(* Logix 5000 project; controller FV vendor 1 type 14 code 217 rev 31.11; software revision 31.00; part 16 of 63 *)
(* tags used below, declared in another part *)
   Dummy : BOOL;
   FR_B230 : INT[255];   // FLOW_BITS Flow Meter Bits
   FR_B240 : INT[255];   // DEBOUNCE Debounce Flags
   FR_B246 : INT[255];   // V_REVERSE Flags for reversing contol action
   FR_B247 : INT[255];   // CHECKWORD Simulation Flags for Checkwords
   FR_B248 : INT[255];   // FORCE ON Force On Flags
   FR_B249 : INT[255];   // FORCE_OFF NOT Force Off Flags
   FR_B3 : INT[255];   // BINARY
   FR_bit_data_file_address : DINT;
   FR_bit_file_bit_offset : DINT;
   FR_bit_file_word_offset : DINT;
   FR_bit_offset : DINT;
   FR_bit_returned : BOOL;
   FR_data_file_value_to_move : DINT;
   FR_from_data_file : DINT;
   FR_from_data_offset : DINT;
   FR_N10 : INT[265];   // FV_AGING Comms to FV Aging PL C
   FR_N100 : INT[265];   // FV FILLING
   FR_N110 : INT[265];   // GREEN BEER Green Beer Main
   FR_N120 : INT[265];   // YEAST CROP Yeast Cropping Main
   FR_N13 : INT[265];   // MV_ROUTE Comms to MV Routing PLC
   FR_N130 : INT[265];   // FILTRATE Filtrate Return
   FR_N14 : INT[265];   // MVFV CIP Comms to MVFV CIP Un it PLC
   FR_N140 : INT[265];   // CIP
   FR_N142 : INT[265];   // CIP
   FR_N143 : INT[265];   // CIP
   FR_N150 : INT[265];   // Original N File From SLC, No Description Available
   FR_N160 : INT[265];   // VESSEL Vessel Working Direc tory
   FR_N170 : INT[265];   // Original N File From SLC, No Description Available
   FR_N180 : INT[265];   // Original N File From SLC, No Description Available
   FR_N198 : INT[265];   // Original N File From SLC, No Description Available
   FR_N20 : INT[265];   // GENERAL General Purpose Setp oints
   FR_N200 : INT[265];   // ANALOG_IN Analog Inputs
   FR_N201 : INT[265];   // Original N File From SLC, No Description Available
   FR_N207 : INT[265];   // Original N File From SLC, No Description Available
   FR_N21 : INT[265];   // CHASE_V FV Filling Beer Chas e Volumes
   FR_N210 : INT[265];   // ANALOG_OUT Analog Outputs
   FR_N220 : INT[265];   // CHECKLIST Checklist Loop Contr ollers
   FR_N225 : INT[265];   // Original N File From SLC, No Description Available
   FR_N226 : INT[265];   // Original N File From SLC, No Description Available
   FR_N245 : INT[265];   // CHECKWORD Checkword Loop Contr ol
   FR_N252 : INT[265];   // OUTPUT_PTR Checkword Pointers t o output flags in B2 50
   FR_N253 : INT[265];   // EN_POINT Pointers to energise d input flags in B25 1
   FR_N254 : INT[265];   // DEN_POINT Pointers to deenergi sed input flags in B 251
   FR_N255 : INT[265];   // CHECKWORDS
   FR_N26 : INT[265];   // FV26
   FR_N27 : INT[265];   // FV27
   FR_N28 : INT[265];   // FV28
   FR_N29 : INT[265];   // FV29
   FR_N30 : INT[265];   // FV30
   FR_N31 : INT[265];   // FV31
   FR_N36 : INT[265];   // Original N File From SLC, No Description Available
   FR_N37 : INT[265];   // Original N File From SLC, No Description Available
   FR_N46 : INT[265];   // Original N File From SLC, No Description Available
   FR_N47 : INT[265];   // Original N File From SLC, No Description Available
   FR_N7 : INT[265];   // INTEGER
   FR_N99 : INT[265];   // COMMENT Comment Lines
   FR_T111 : TIMER[255];   // GREEN BEER
(* FR_Common, continued *)

ROUTINE FR_Get_NFile_Value   (* ladder *)
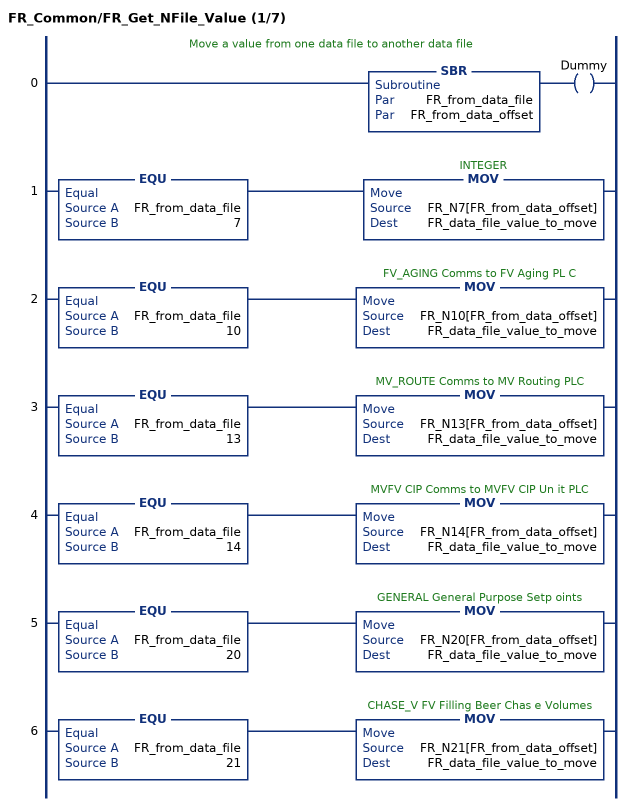
   // Move a value from one data file to another data file
   0: SBR(FR_from_data_file,FR_from_data_offset)OTE(Dummy);
   1: EQU(FR_from_data_file,7)MOV(FR_N7[FR_from_data_offset],FR_data_file_value_to_move);
   2: EQU(FR_from_data_file,10)MOV(FR_N10[FR_from_data_offset],FR_data_file_value_to_move);
   3: EQU(FR_from_data_file,13)MOV(FR_N13[FR_from_data_offset],FR_data_file_value_to_move);
   4: EQU(FR_from_data_file,14)MOV(FR_N14[FR_from_data_offset],FR_data_file_value_to_move);
   5: EQU(FR_from_data_file,20)MOV(FR_N20[FR_from_data_offset],FR_data_file_value_to_move);
   6: EQU(FR_from_data_file,21)MOV(FR_N21[FR_from_data_offset],FR_data_file_value_to_move);
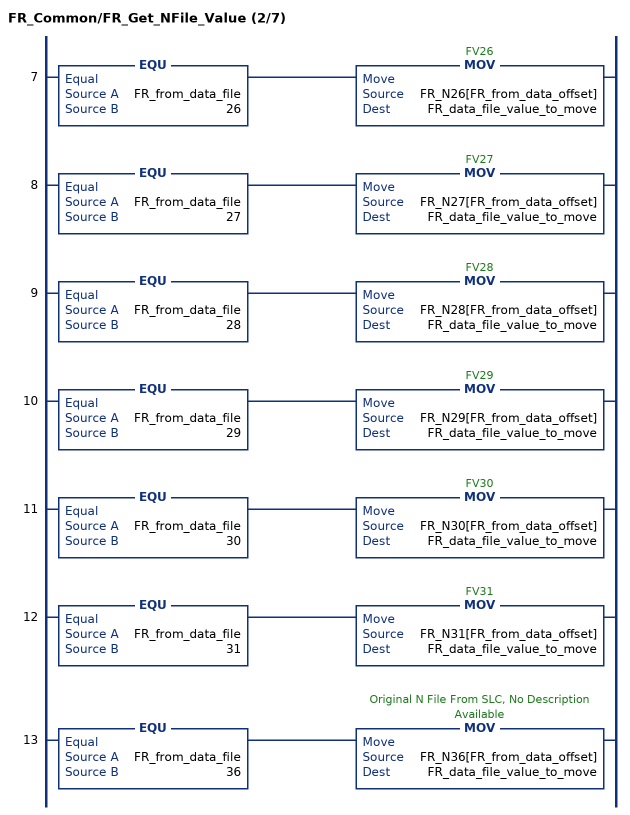
   7: EQU(FR_from_data_file,26)MOV(FR_N26[FR_from_data_offset],FR_data_file_value_to_move);
   8: EQU(FR_from_data_file,27)MOV(FR_N27[FR_from_data_offset],FR_data_file_value_to_move);
   9: EQU(FR_from_data_file,28)MOV(FR_N28[FR_from_data_offset],FR_data_file_value_to_move);
   10: EQU(FR_from_data_file,29)MOV(FR_N29[FR_from_data_offset],FR_data_file_value_to_move);
   11: EQU(FR_from_data_file,30)MOV(FR_N30[FR_from_data_offset],FR_data_file_value_to_move);
   12: EQU(FR_from_data_file,31)MOV(FR_N31[FR_from_data_offset],FR_data_file_value_to_move);
   13: EQU(FR_from_data_file,36)MOV(FR_N36[FR_from_data_offset],FR_data_file_value_to_move);
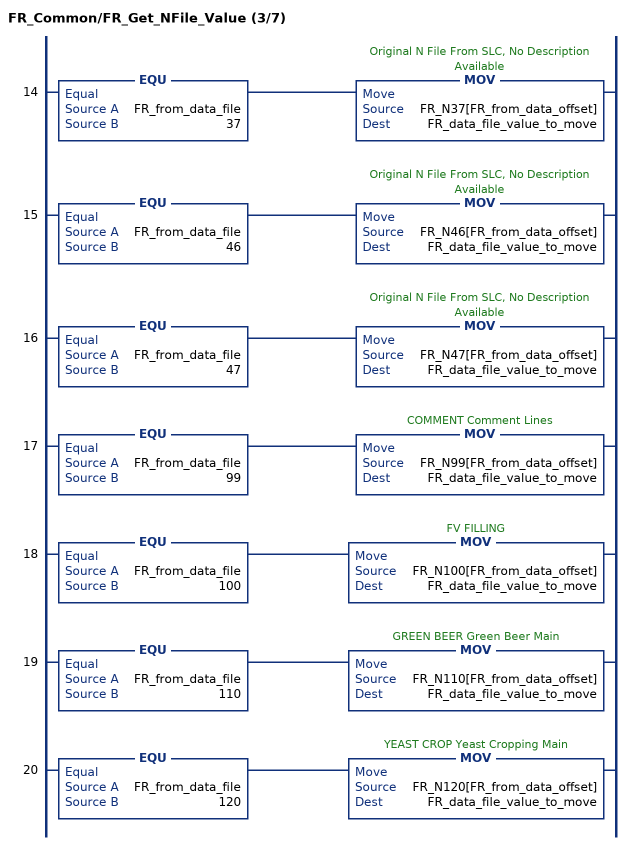
   14: EQU(FR_from_data_file,37)MOV(FR_N37[FR_from_data_offset],FR_data_file_value_to_move);
   15: EQU(FR_from_data_file,46)MOV(FR_N46[FR_from_data_offset],FR_data_file_value_to_move);
   16: EQU(FR_from_data_file,47)MOV(FR_N47[FR_from_data_offset],FR_data_file_value_to_move);
   17: EQU(FR_from_data_file,99)MOV(FR_N99[FR_from_data_offset],FR_data_file_value_to_move);
   18: EQU(FR_from_data_file,100)MOV(FR_N100[FR_from_data_offset],FR_data_file_value_to_move);
   19: EQU(FR_from_data_file,110)MOV(FR_N110[FR_from_data_offset],FR_data_file_value_to_move);
   20: EQU(FR_from_data_file,120)MOV(FR_N120[FR_from_data_offset],FR_data_file_value_to_move);
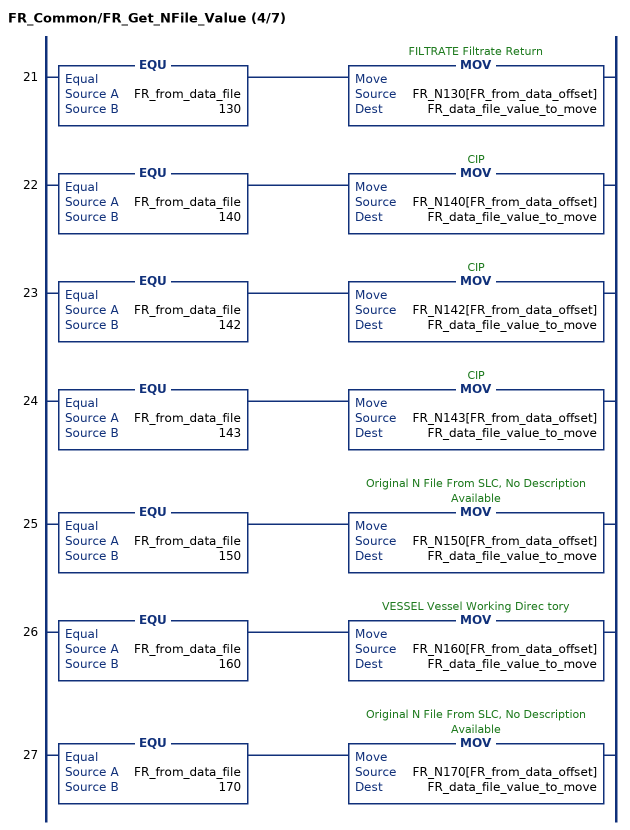
   21: EQU(FR_from_data_file,130)MOV(FR_N130[FR_from_data_offset],FR_data_file_value_to_move);
   22: EQU(FR_from_data_file,140)MOV(FR_N140[FR_from_data_offset],FR_data_file_value_to_move);
   23: EQU(FR_from_data_file,142)MOV(FR_N142[FR_from_data_offset],FR_data_file_value_to_move);
   24: EQU(FR_from_data_file,143)MOV(FR_N143[FR_from_data_offset],FR_data_file_value_to_move);
   25: EQU(FR_from_data_file,150)MOV(FR_N150[FR_from_data_offset],FR_data_file_value_to_move);
   26: EQU(FR_from_data_file,160)MOV(FR_N160[FR_from_data_offset],FR_data_file_value_to_move);
   27: EQU(FR_from_data_file,170)MOV(FR_N170[FR_from_data_offset],FR_data_file_value_to_move);
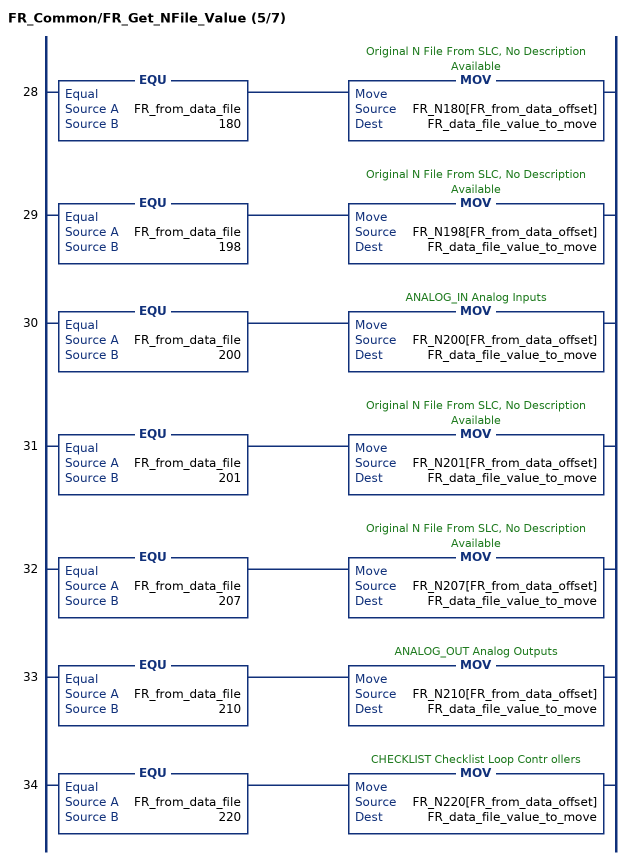
   28: EQU(FR_from_data_file,180)MOV(FR_N180[FR_from_data_offset],FR_data_file_value_to_move);
   29: EQU(FR_from_data_file,198)MOV(FR_N198[FR_from_data_offset],FR_data_file_value_to_move);
   30: EQU(FR_from_data_file,200)MOV(FR_N200[FR_from_data_offset],FR_data_file_value_to_move);
   31: EQU(FR_from_data_file,201)MOV(FR_N201[FR_from_data_offset],FR_data_file_value_to_move);
   32: EQU(FR_from_data_file,207)MOV(FR_N207[FR_from_data_offset],FR_data_file_value_to_move);
   33: EQU(FR_from_data_file,210)MOV(FR_N210[FR_from_data_offset],FR_data_file_value_to_move);
   34: EQU(FR_from_data_file,220)MOV(FR_N220[FR_from_data_offset],FR_data_file_value_to_move);
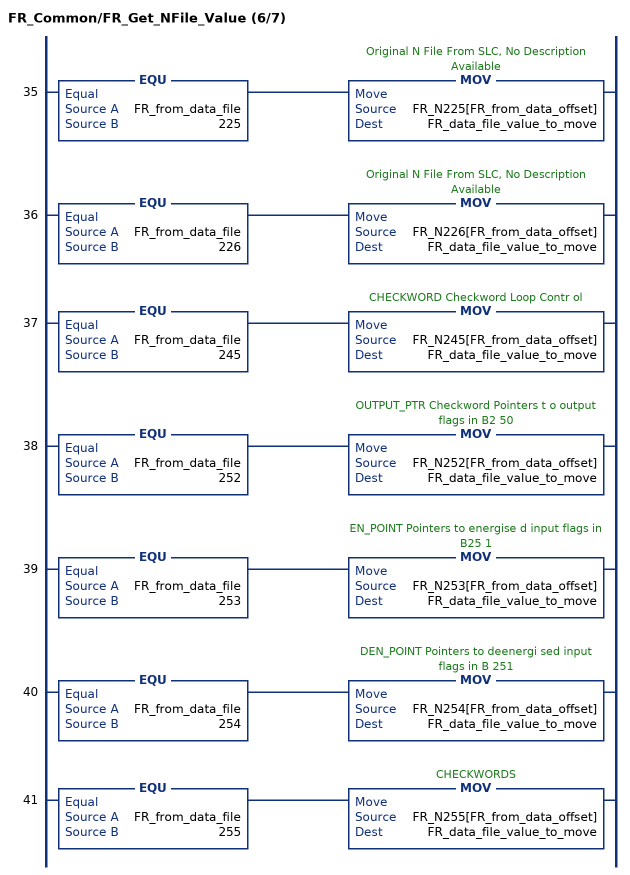
   35: EQU(FR_from_data_file,225)MOV(FR_N225[FR_from_data_offset],FR_data_file_value_to_move);
   36: EQU(FR_from_data_file,226)MOV(FR_N226[FR_from_data_offset],FR_data_file_value_to_move);
   37: EQU(FR_from_data_file,245)MOV(FR_N245[FR_from_data_offset],FR_data_file_value_to_move);
   38: EQU(FR_from_data_file,252)MOV(FR_N252[FR_from_data_offset],FR_data_file_value_to_move);
   39: EQU(FR_from_data_file,253)MOV(FR_N253[FR_from_data_offset],FR_data_file_value_to_move);
   40: EQU(FR_from_data_file,254)MOV(FR_N254[FR_from_data_offset],FR_data_file_value_to_move);
   41: EQU(FR_from_data_file,255)MOV(FR_N255[FR_from_data_offset],FR_data_file_value_to_move);
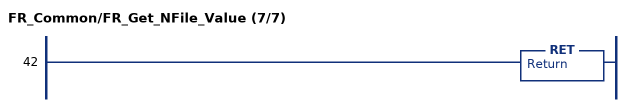
   42: RET();
END_ROUTINE

ROUTINE FR_GetBitFile_Value   (* ladder *)
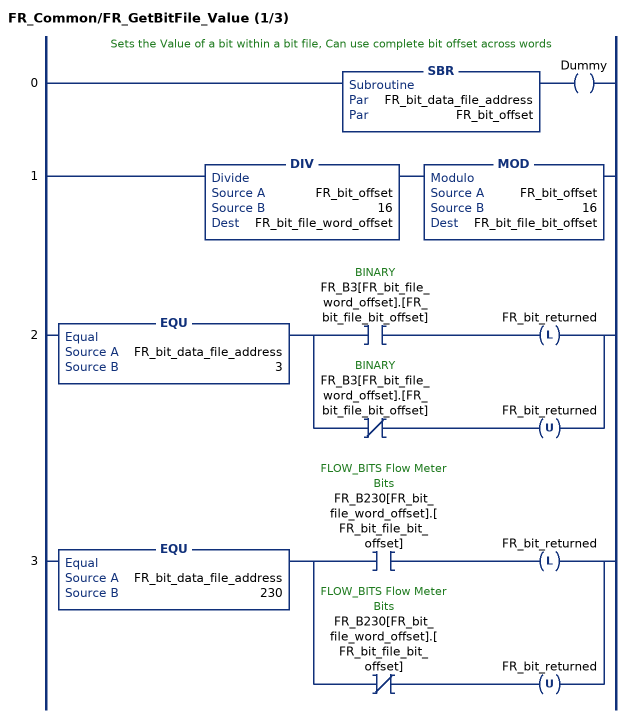
   // Sets the Value of a bit within a bit file, Can use complete bit offset across words
   0: SBR(FR_bit_data_file_address,FR_bit_offset)OTE(Dummy);
   1: DIV(FR_bit_offset,16,FR_bit_file_word_offset)MOD(FR_bit_offset,16,FR_bit_file_bit_offset);
   2: EQU(FR_bit_data_file_address,3)[XIC(FR_B3[FR_bit_file_word_offset].[FR_bit_file_bit_offset]) OTL(FR_bit_returned) ,XIO(FR_B3[FR_bit_file_word_offset].[FR_bit_file_bit_offset]) OTU(FR_bit_returned) ];
   3: EQU(FR_bit_data_file_address,230)[XIC(FR_B230[FR_bit_file_word_offset].[FR_bit_file_bit_offset]) OTL(FR_bit_returned) ,XIO(FR_B230[FR_bit_file_word_offset].[FR_bit_file_bit_offset]) OTU(FR_bit_returned) ];
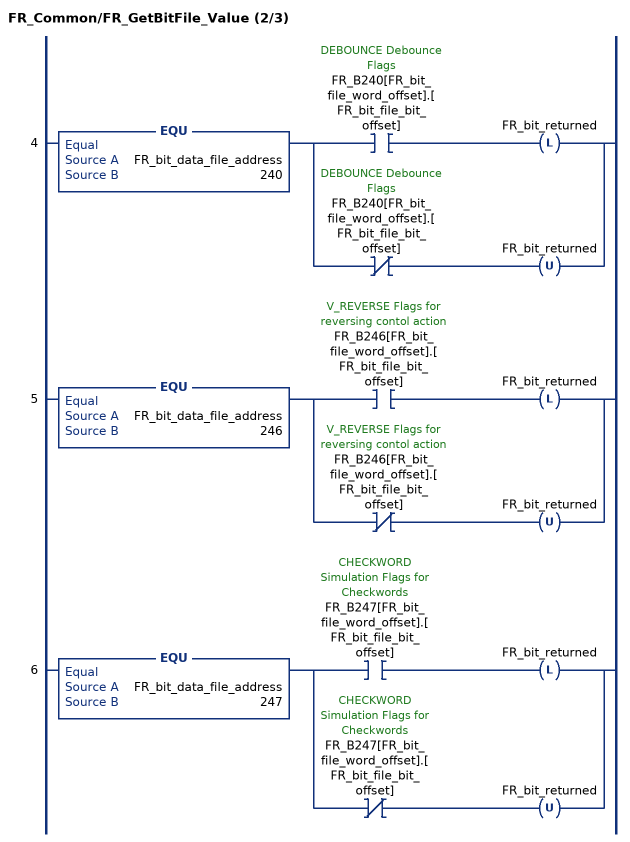
   4: EQU(FR_bit_data_file_address,240)[XIC(FR_B240[FR_bit_file_word_offset].[FR_bit_file_bit_offset]) OTL(FR_bit_returned) ,XIO(FR_B240[FR_bit_file_word_offset].[FR_bit_file_bit_offset]) OTU(FR_bit_returned) ];
   5: EQU(FR_bit_data_file_address,246)[XIC(FR_B246[FR_bit_file_word_offset].[FR_bit_file_bit_offset]) OTL(FR_bit_returned) ,XIO(FR_B246[FR_bit_file_word_offset].[FR_bit_file_bit_offset]) OTU(FR_bit_returned) ];
   6: EQU(FR_bit_data_file_address,247)[XIC(FR_B247[FR_bit_file_word_offset].[FR_bit_file_bit_offset]) OTL(FR_bit_returned) ,XIO(FR_B247[FR_bit_file_word_offset].[FR_bit_file_bit_offset]) OTU(FR_bit_returned) ];
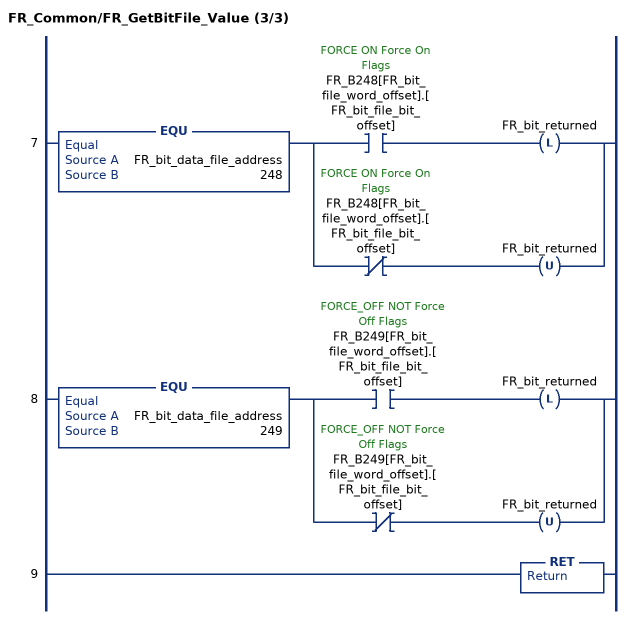
   7: EQU(FR_bit_data_file_address,248)[XIC(FR_B248[FR_bit_file_word_offset].[FR_bit_file_bit_offset]) OTL(FR_bit_returned) ,XIO(FR_B248[FR_bit_file_word_offset].[FR_bit_file_bit_offset]) OTU(FR_bit_returned) ];
   8: EQU(FR_bit_data_file_address,249)[XIC(FR_B249[FR_bit_file_word_offset].[FR_bit_file_bit_offset]) OTL(FR_bit_returned) ,XIO(FR_B249[FR_bit_file_word_offset].[FR_bit_file_bit_offset]) OTU(FR_bit_returned) ];
   9: RET();
END_ROUTINE

ROUTINE FR_GRN_BEER_111   (* ladder *)
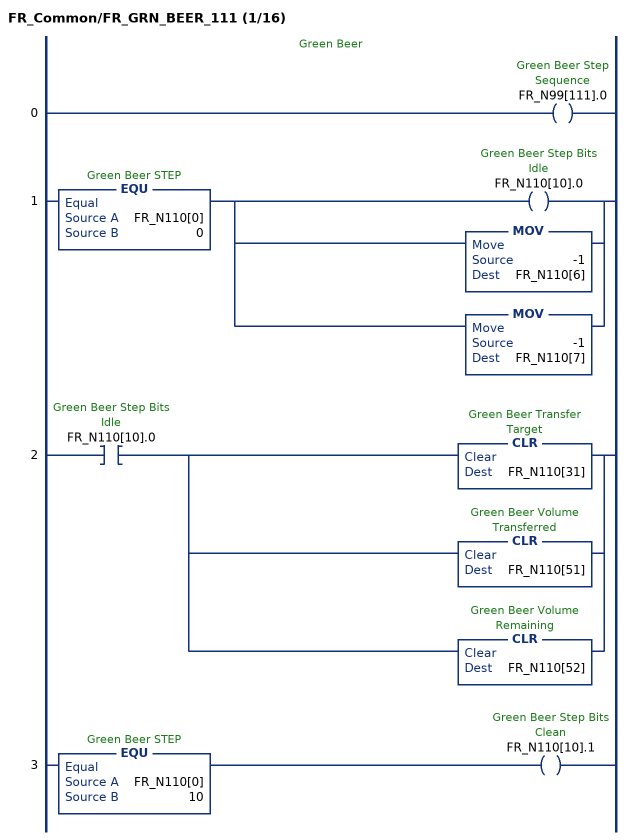
   // Green Beer
   0: OTE(FR_N99[111].0);
   1: EQU(FR_N110[0],0)[OTE(FR_N110[10].0) ,MOV(-1,FR_N110[6]) ,MOV(-1,FR_N110[7]) ];
   2: XIC(FR_N110[10].0)[CLR(FR_N110[31]) ,CLR(FR_N110[51]) ,CLR(FR_N110[52]) ];
   3: EQU(FR_N110[0],10)OTE(FR_N110[10].1);
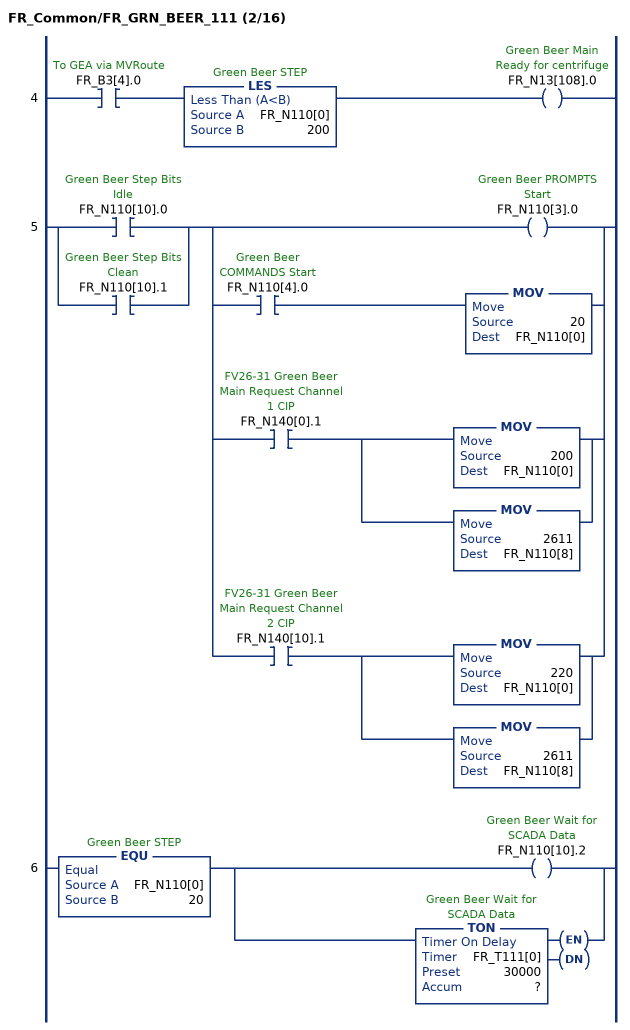
   4: XIC(FR_B3[4].0)LES(FR_N110[0],200)OTE(FR_N13[108].0);
   5: [XIC(FR_N110[10].0) ,XIC(FR_N110[10].1) ][OTE(FR_N110[3].0) ,XIC(FR_N110[4].0) MOV(20,FR_N110[0]) ,XIC(FR_N140[0].1) [MOV(200,FR_N110[0]) ,MOV(2611,FR_N110[8]) ] ,XIC(FR_N140[10].1) [MOV(220,FR_N110[0]) ,MOV(2611,FR_N110[8]) ] ];
   6: EQU(FR_N110[0],20)[OTE(FR_N110[10].2) ,TON(FR_T111[0],?,?) ];
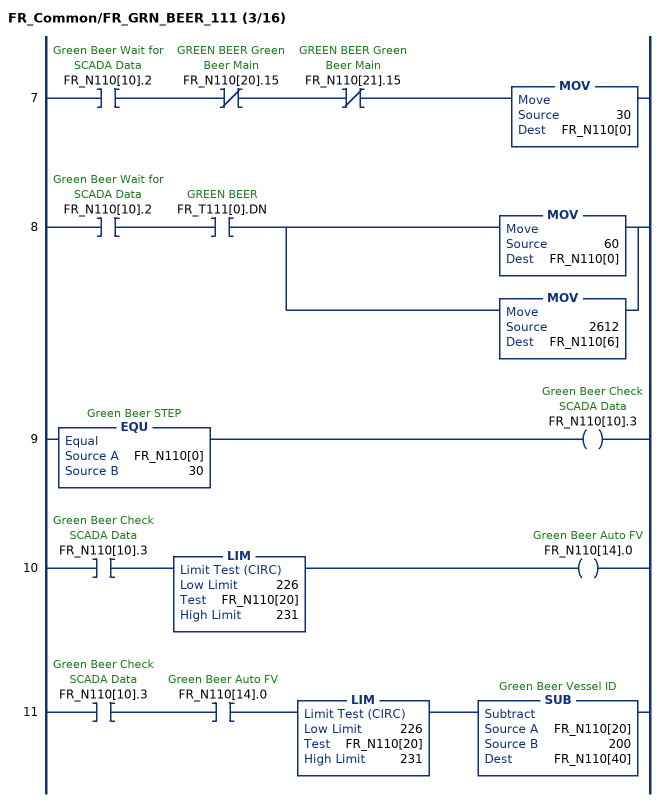
   7: XIC(FR_N110[10].2)XIO(FR_N110[20].15)XIO(FR_N110[21].15)MOV(30,FR_N110[0]);
   8: XIC(FR_N110[10].2)XIC(FR_T111[0].DN)[MOV(60,FR_N110[0]) ,MOV(2612,FR_N110[6]) ];
   9: EQU(FR_N110[0],30)OTE(FR_N110[10].3);
   10: XIC(FR_N110[10].3)LIM(226,FR_N110[20],231)OTE(FR_N110[14].0);
   11: XIC(FR_N110[10].3)XIC(FR_N110[14].0)LIM(226,FR_N110[20],231)SUB(FR_N110[20],200,FR_N110[40]);
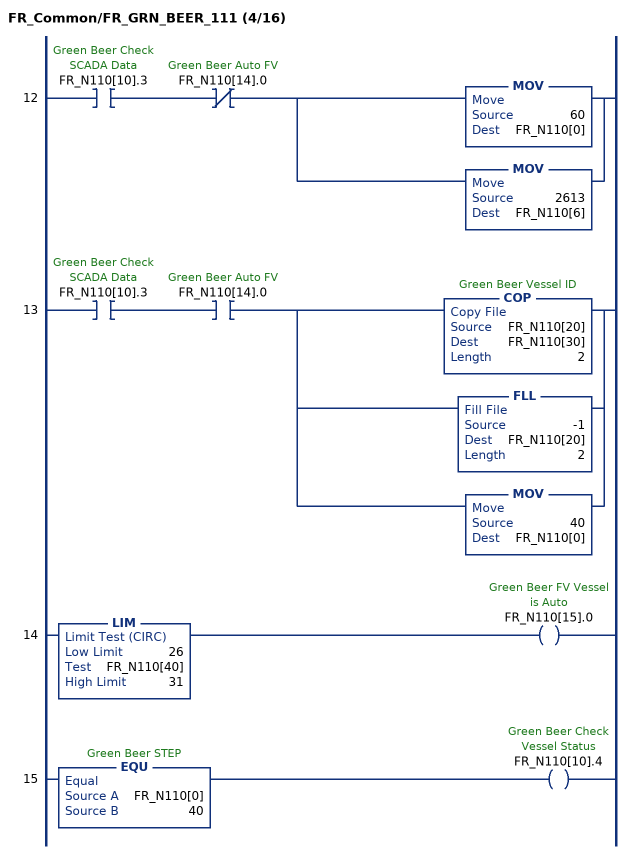
   12: XIC(FR_N110[10].3)XIO(FR_N110[14].0)[MOV(60,FR_N110[0]) ,MOV(2613,FR_N110[6]) ];
   13: XIC(FR_N110[10].3)XIC(FR_N110[14].0)[COP(FR_N110[20],FR_N110[30],2) ,FLL(-1,FR_N110[20],2) ,MOV(40,FR_N110[0]) ];
   14: LIM(26,FR_N110[40],31)OTE(FR_N110[15].0);
   15: EQU(FR_N110[0],40)OTE(FR_N110[10].4);
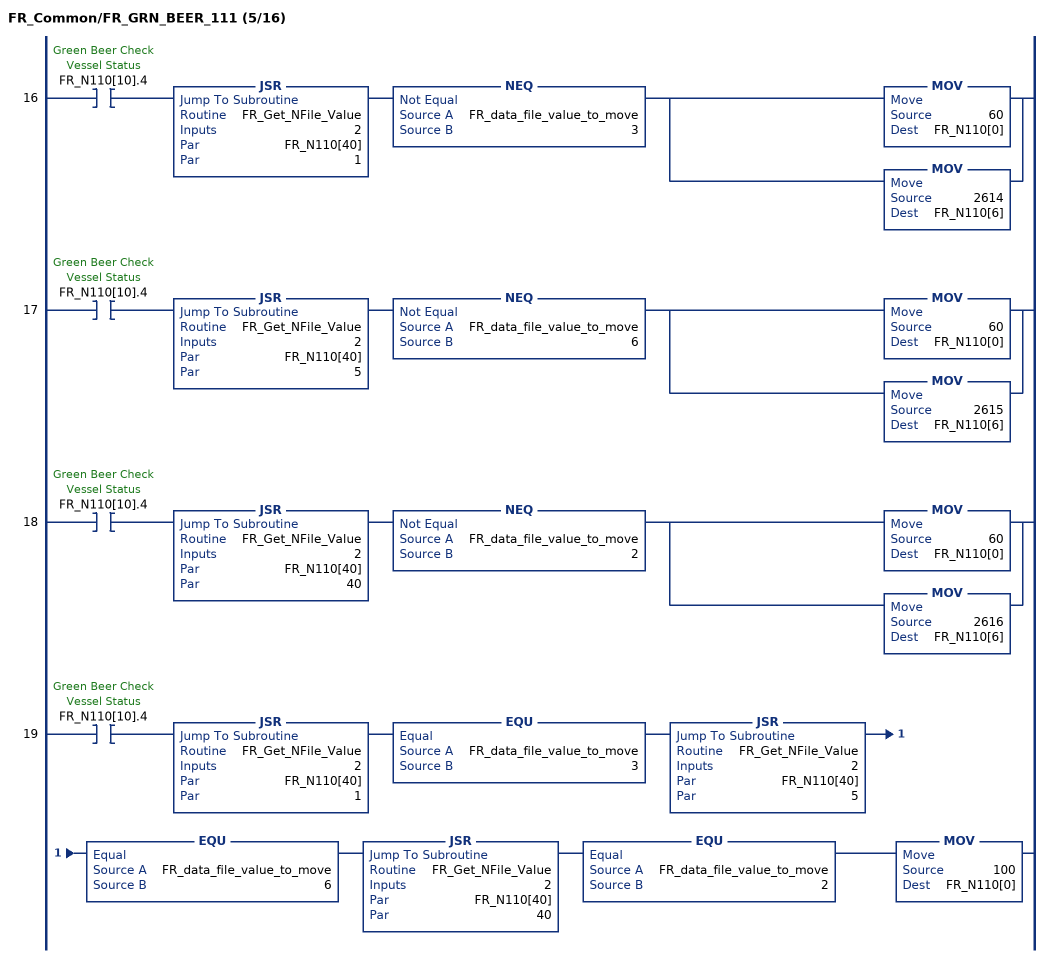
   16: XIC(FR_N110[10].4)JSR(FR_Get_NFile_Value,2,FR_N110[40],1)NEQ(FR_data_file_value_to_move,3)[MOV(60,FR_N110[0]) ,MOV(2614,FR_N110[6]) ];
   17: XIC(FR_N110[10].4)JSR(FR_Get_NFile_Value,2,FR_N110[40],5)NEQ(FR_data_file_value_to_move,6)[MOV(60,FR_N110[0]) ,MOV(2615,FR_N110[6]) ];
   18: XIC(FR_N110[10].4)JSR(FR_Get_NFile_Value,2,FR_N110[40],40)NEQ(FR_data_file_value_to_move,2)[MOV(60,FR_N110[0]) ,MOV(2616,FR_N110[6]) ];
   19: XIC(FR_N110[10].4)JSR(FR_Get_NFile_Value,2,FR_N110[40],1)EQU(FR_data_file_value_to_move,3)JSR(FR_Get_NFile_Value,2,FR_N110[40],5)EQU(FR_data_file_value_to_move,6)JSR(FR_Get_NFile_Value,2,FR_N110[40],40)EQU(FR_data_file_value_to_move,2)MOV(100,FR_N110[0]);
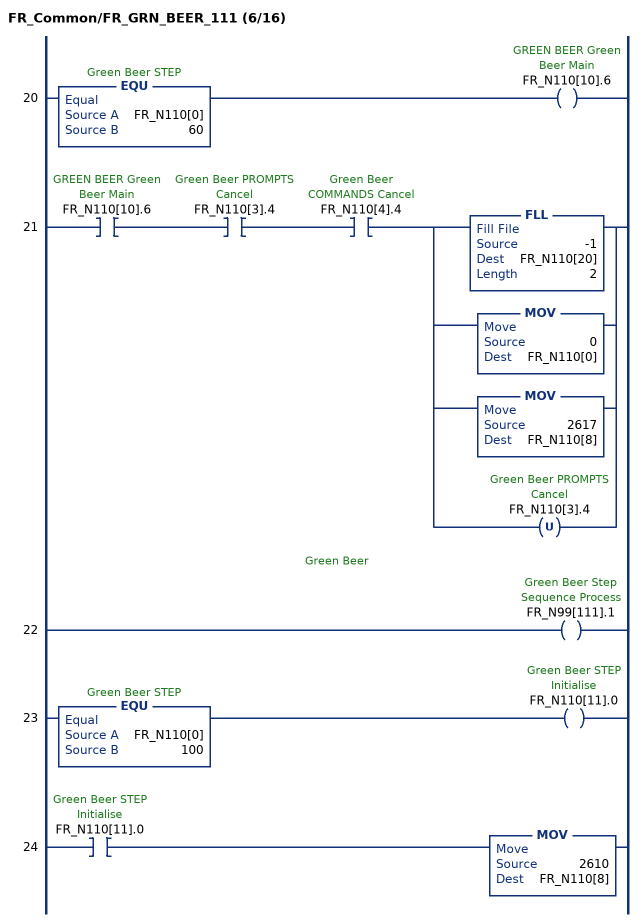
   20: EQU(FR_N110[0],60)OTE(FR_N110[10].6);
   21: XIC(FR_N110[10].6)XIC(FR_N110[3].4)XIC(FR_N110[4].4)[FLL(-1,FR_N110[20],2) ,MOV(0,FR_N110[0]) ,MOV(2617,FR_N110[8]) ,OTU(FR_N110[3].4) ];
   // Green Beer
   22: OTE(FR_N99[111].1);
   23: EQU(FR_N110[0],100)OTE(FR_N110[11].0);
   24: XIC(FR_N110[11].0)MOV(2610,FR_N110[8]);
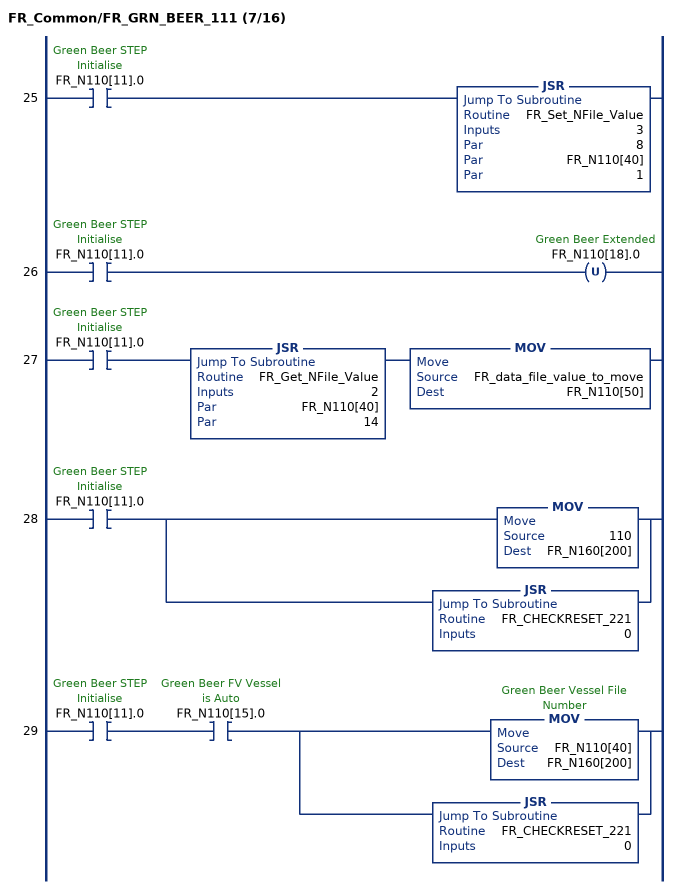
   25: XIC(FR_N110[11].0)JSR(FR_Set_NFile_Value,3,8,FR_N110[40],1);
   26: XIC(FR_N110[11].0)OTU(FR_N110[18].0);
   27: XIC(FR_N110[11].0)JSR(FR_Get_NFile_Value,2,FR_N110[40],14)MOV(FR_data_file_value_to_move,FR_N110[50]);
   28: XIC(FR_N110[11].0)[MOV(110,FR_N160[200]) ,JSR(FR_CHECKRESET_221,0) ];
   29: XIC(FR_N110[11].0)XIC(FR_N110[15].0)[MOV(FR_N110[40],FR_N160[200]) ,JSR(FR_CHECKRESET_221,0) ];
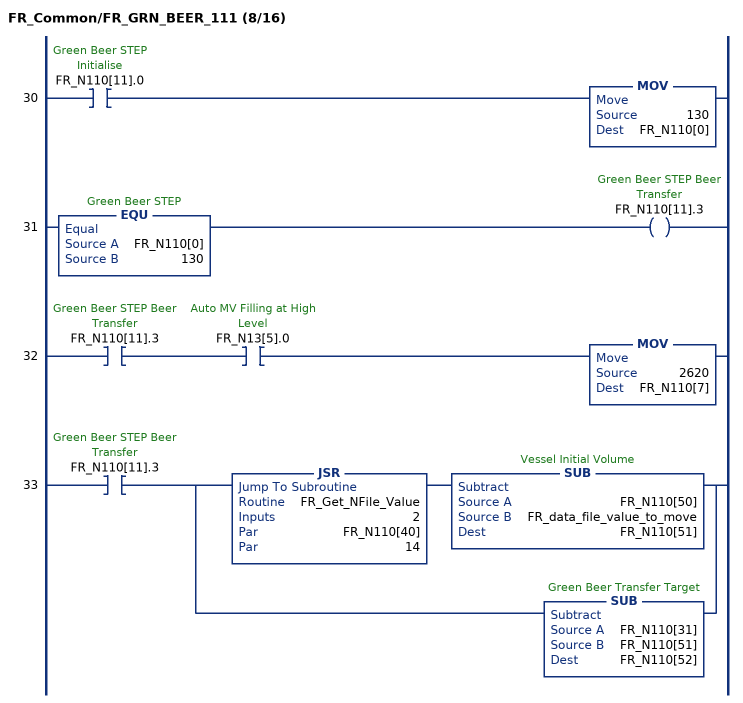
   30: XIC(FR_N110[11].0)MOV(130,FR_N110[0]);
   31: EQU(FR_N110[0],130)OTE(FR_N110[11].3);
   32: XIC(FR_N110[11].3)XIC(FR_N13[5].0)MOV(2620,FR_N110[7]);
   33: XIC(FR_N110[11].3)[JSR(FR_Get_NFile_Value,2,FR_N110[40],14) SUB(FR_N110[50],FR_data_file_value_to_move,FR_N110[51]) ,SUB(FR_N110[31],FR_N110[51],FR_N110[52]) ];
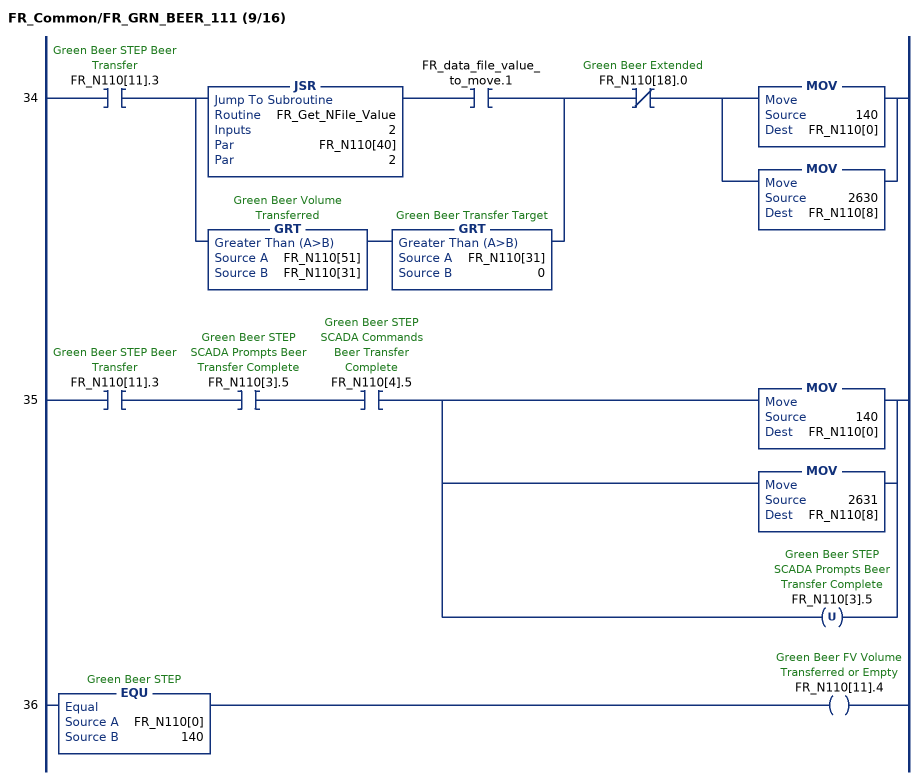
   34: XIC(FR_N110[11].3)[JSR(FR_Get_NFile_Value,2,FR_N110[40],2) XIC(FR_data_file_value_to_move.1) ,GRT(FR_N110[51],FR_N110[31]) GRT(FR_N110[31],0) ]XIO(FR_N110[18].0)[MOV(140,FR_N110[0]) ,MOV(2630,FR_N110[8]) ];
   35: XIC(FR_N110[11].3)XIC(FR_N110[3].5)XIC(FR_N110[4].5)[MOV(140,FR_N110[0]) ,MOV(2631,FR_N110[8]) ,OTU(FR_N110[3].5) ];
   36: EQU(FR_N110[0],140)OTE(FR_N110[11].4);
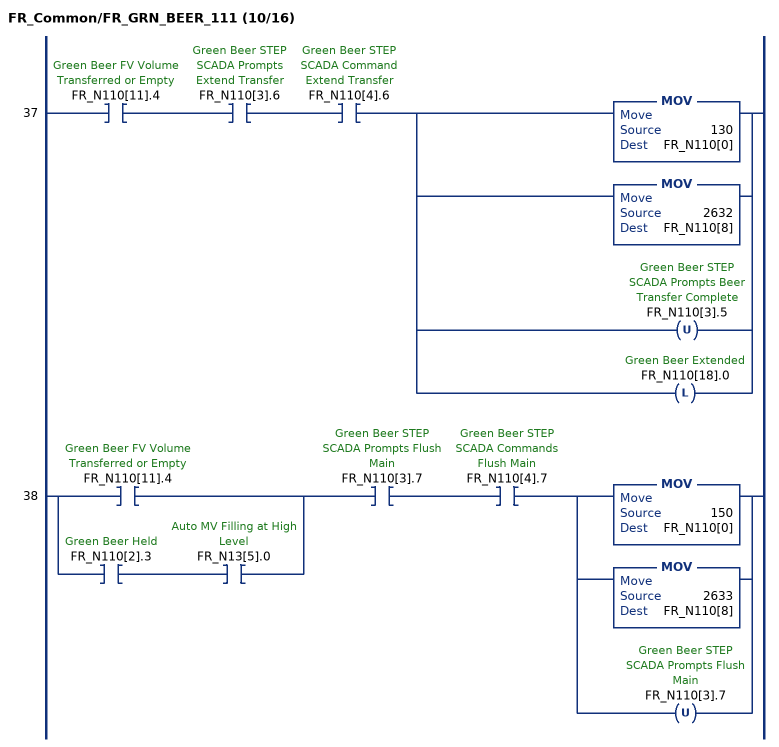
   37: XIC(FR_N110[11].4)XIC(FR_N110[3].6)XIC(FR_N110[4].6)[MOV(130,FR_N110[0]) ,MOV(2632,FR_N110[8]) ,OTU(FR_N110[3].5) ,OTL(FR_N110[18].0) ];
   38: [XIC(FR_N110[11].4) ,XIC(FR_N110[2].3) XIC(FR_N13[5].0) ]XIC(FR_N110[3].7)XIC(FR_N110[4].7)[MOV(150,FR_N110[0]) ,MOV(2633,FR_N110[8]) ,OTU(FR_N110[3].7) ];
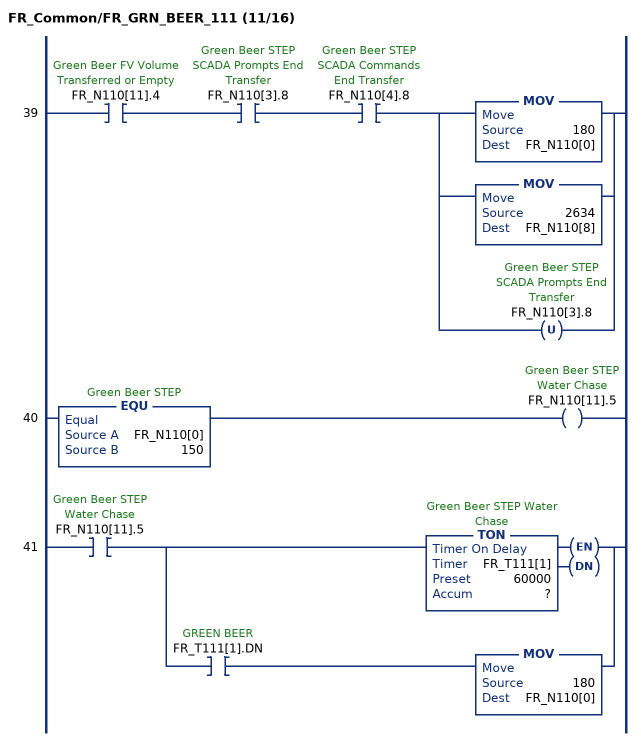
   39: XIC(FR_N110[11].4)XIC(FR_N110[3].8)XIC(FR_N110[4].8)[MOV(180,FR_N110[0]) ,MOV(2634,FR_N110[8]) ,OTU(FR_N110[3].8) ];
   40: EQU(FR_N110[0],150)OTE(FR_N110[11].5);
   41: XIC(FR_N110[11].5)[TON(FR_T111[1],?,?) ,XIC(FR_T111[1].DN) MOV(180,FR_N110[0]) ];
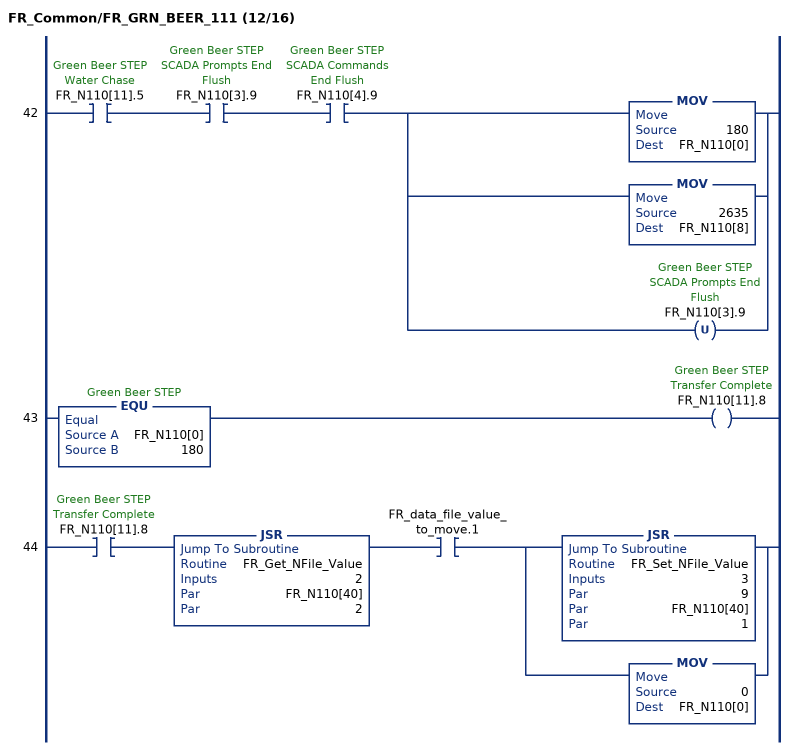
   42: XIC(FR_N110[11].5)XIC(FR_N110[3].9)XIC(FR_N110[4].9)[MOV(180,FR_N110[0]) ,MOV(2635,FR_N110[8]) ,OTU(FR_N110[3].9) ];
   43: EQU(FR_N110[0],180)OTE(FR_N110[11].8);
   44: XIC(FR_N110[11].8)JSR(FR_Get_NFile_Value,2,FR_N110[40],2)XIC(FR_data_file_value_to_move.1)[JSR(FR_Set_NFile_Value,3,9,FR_N110[40],1) ,MOV(0,FR_N110[0]) ];
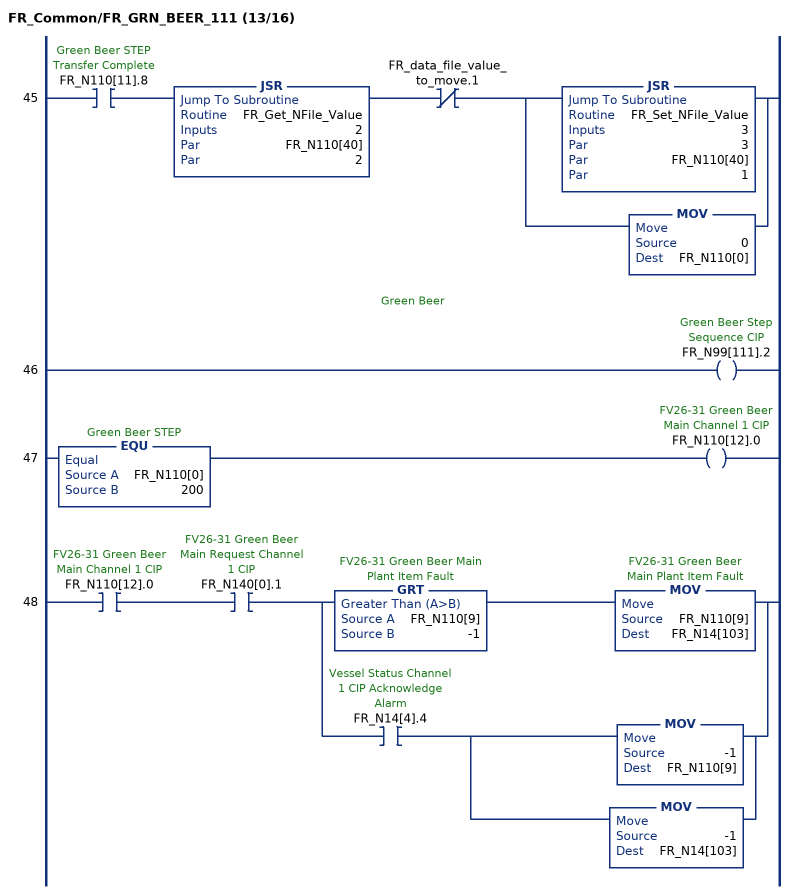
   45: XIC(FR_N110[11].8)JSR(FR_Get_NFile_Value,2,FR_N110[40],2)XIO(FR_data_file_value_to_move.1)[JSR(FR_Set_NFile_Value,3,3,FR_N110[40],1) ,MOV(0,FR_N110[0]) ];
   // Green Beer
   46: OTE(FR_N99[111].2);
   47: EQU(FR_N110[0],200)OTE(FR_N110[12].0);
   48: XIC(FR_N110[12].0)XIC(FR_N140[0].1)[GRT(FR_N110[9],-1) MOV(FR_N110[9],FR_N14[103]) ,XIC(FR_N14[4].4) [MOV(-1,FR_N110[9]) ,MOV(-1,FR_N14[103]) ] ];
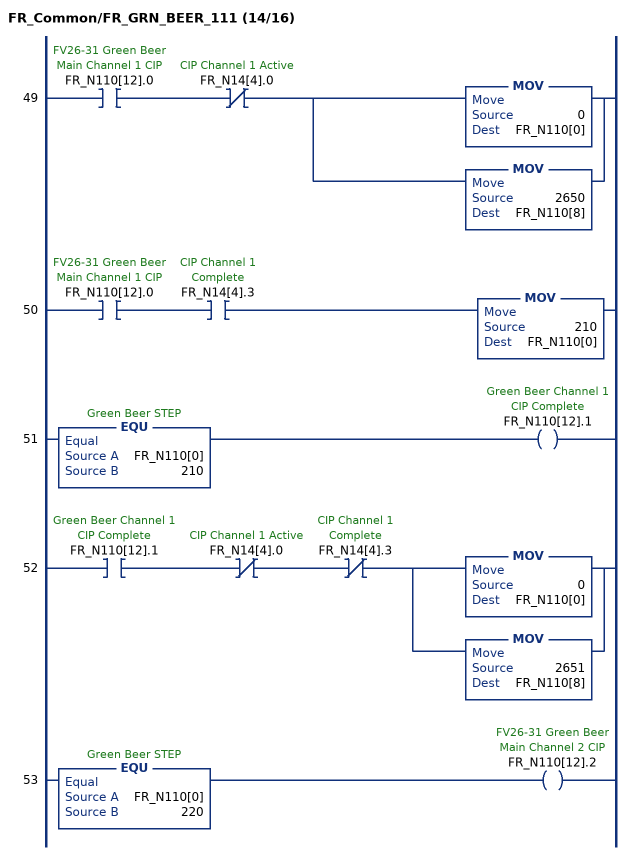
   49: XIC(FR_N110[12].0)XIO(FR_N14[4].0)[MOV(0,FR_N110[0]) ,MOV(2650,FR_N110[8]) ];
   50: XIC(FR_N110[12].0)XIC(FR_N14[4].3)MOV(210,FR_N110[0]);
   51: EQU(FR_N110[0],210)OTE(FR_N110[12].1);
   52: XIC(FR_N110[12].1)XIO(FR_N14[4].0)XIO(FR_N14[4].3)[MOV(0,FR_N110[0]) ,MOV(2651,FR_N110[8]) ];
   53: EQU(FR_N110[0],220)OTE(FR_N110[12].2);
